   		COP(N746[TMP_dSourceOffset], N14[TMP_dDestOffset], TMP_dNumValues);
   	ELSIF (TMP_dSourceFile = 747) AND (TMP_dDestFile = 14) THEN
   		COP(N747[TMP_dSourceOffset], N14[TMP_dDestOffset], TMP_dNumValues);
   	ELSIF (TMP_dSourceFile = 748) AND (TMP_dDestFile = 14) THEN
   		COP(N748[TMP_dSourceOffset], N14[TMP_dDestOffset], TMP_dNumValues);
   	ELSIF (TMP_dSourceFile = 749) AND (TMP_dDestFile = 14) THEN
   		COP(N749[TMP_dSourceOffset], N14[TMP_dDestOffset], TMP_dNumValues);
   	ELSIF (TMP_dSourceFile = 750) AND (TMP_dDestFile = 14) THEN
   		COP(N750[TMP_dSourceOffset], N14[TMP_dDestOffset], TMP_dNumValues);
   	ELSIF (TMP_dSourceFile = 751) AND (TMP_dDestFile = 14) THEN
   		COP(N751[TMP_dSourceOffset], N14[TMP_dDestOffset], TMP_dNumValues);
   	ELSIF (TMP_dSourceFile = 752) AND (TMP_dDestFile = 14) THEN
   		COP(N752[TMP_dSourceOffset], N14[TMP_dDestOffset], TMP_dNumValues);
   	ELSIF (TMP_dSourceFile = 753) AND (TMP_dDestFile = 14) THEN
   		COP(N753[TMP_dSourceOffset], N14[TMP_dDestOffset], TMP_dNumValues);
   	ELSIF (TMP_dSourceFile = 754) AND (TMP_dDestFile = 14) THEN
   		COP(N754[TMP_dSourceOffset], N14[TMP_dDestOffset], TMP_dNumValues);
   	ELSIF (TMP_dSourceFile = 755) AND (TMP_dDestFile = 14) THEN
   		COP(N755[TMP_dSourceOffset], N14[TMP_dDestOffset], TMP_dNumValues);
   	ELSIF (TMP_dSourceFile = 756) AND (TMP_dDestFile = 14) THEN
   		COP(N756[TMP_dSourceOffset], N14[TMP_dDestOffset], TMP_dNumValues);
   	ELSIF (TMP_dSourceFile = 757) AND (TMP_dDestFile = 14) THEN
   		COP(N757[TMP_dSourceOffset], N14[TMP_dDestOffset], TMP_dNumValues);
   	ELSIF (TMP_dSourceFile = 758) AND (TMP_dDestFile = 14) THEN
   		COP(N758[TMP_dSourceOffset], N14[TMP_dDestOffset], TMP_dNumValues);
   	ELSIF (TMP_dSourceFile = 759) AND (TMP_dDestFile = 14) THEN
   		COP(N759[TMP_dSourceOffset], N14[TMP_dDestOffset], TMP_dNumValues);
   	ELSIF (TMP_dSourceFile = 760) AND (TMP_dDestFile = 14) THEN
   		COP(N760[TMP_dSourceOffset], N14[TMP_dDestOffset], TMP_dNumValues);
   	ELSIF (TMP_dSourceFile = 761) AND (TMP_dDestFile = 14) THEN
   		COP(N761[TMP_dSourceOffset], N14[TMP_dDestOffset], TMP_dNumValues);
   	ELSIF (TMP_dSourceFile = 762) AND (TMP_dDestFile = 14) THEN
   		COP(N762[TMP_dSourceOffset], N14[TMP_dDestOffset], TMP_dNumValues);
   	ELSIF (TMP_dSourceFile = 763) AND (TMP_dDestFile = 14) THEN
   		COP(N763[TMP_dSourceOffset], N14[TMP_dDestOffset], TMP_dNumValues);
   	ELSIF (TMP_dSourceFile = 764) AND (TMP_dDestFile = 14) THEN
   		COP(N764[TMP_dSourceOffset], N14[TMP_dDestOffset], TMP_dNumValues);
   	ELSIF (TMP_dSourceFile = 765) AND (TMP_dDestFile = 14) THEN
   		COP(N765[TMP_dSourceOffset], N14[TMP_dDestOffset], TMP_dNumValues);
   	ELSIF (TMP_dSourceFile = 766) AND (TMP_dDestFile = 14) THEN
   		COP(N766[TMP_dSourceOffset], N14[TMP_dDestOffset], TMP_dNumValues);
   	ELSIF (TMP_dSourceFile = 767) AND (TMP_dDestFile = 14) THEN
   		COP(N767[TMP_dSourceOffset], N14[TMP_dDestOffset], TMP_dNumValues);
   	ELSIF (TMP_dSourceFile = 768) AND (TMP_dDestFile = 14) THEN
   		COP(N768[TMP_dSourceOffset], N14[TMP_dDestOffset], TMP_dNumValues);
   	ELSIF (TMP_dSourceFile = 769) AND (TMP_dDestFile = 14) THEN
   		COP(N769[TMP_dSourceOffset], N14[TMP_dDestOffset], TMP_dNumValues);
   	ELSIF (TMP_dSourceFile = 770) AND (TMP_dDestFile = 14) THEN
   		COP(N770[TMP_dSourceOffset], N14[TMP_dDestOffset], TMP_dNumValues);
   	ELSIF (TMP_dSourceFile = 771) AND (TMP_dDestFile = 14) THEN
   		COP(N771[TMP_dSourceOffset], N14[TMP_dDestOffset], TMP_dNumValues);
   	ELSIF (TMP_dSourceFile = 772) AND (TMP_dDestFile = 14) THEN
   		COP(N772[TMP_dSourceOffset], N14[TMP_dDestOffset], TMP_dNumValues);
   	ELSIF (TMP_dSourceFile = 773) AND (TMP_dDestFile = 14) THEN
   		COP(N773[TMP_dSourceOffset], N14[TMP_dDestOffset], TMP_dNumValues);
   	ELSIF (TMP_dSourceFile = 774) AND (TMP_dDestFile = 14) THEN
   		COP(N774[TMP_dSourceOffset], N14[TMP_dDestOffset], TMP_dNumValues);
   	ELSIF (TMP_dSourceFile = 775) AND (TMP_dDestFile = 14) THEN
   		COP(N775[TMP_dSourceOffset], N14[TMP_dDestOffset], TMP_dNumValues);
   	ELSIF (TMP_dSourceFile = 776) AND (TMP_dDestFile = 14) THEN
   		COP(N776[TMP_dSourceOffset], N14[TMP_dDestOffset], TMP_dNumValues);
   	ELSIF (TMP_dSourceFile = 777) AND (TMP_dDestFile = 14) THEN
   		COP(N777[TMP_dSourceOffset], N14[TMP_dDestOffset], TMP_dNumValues);
   	ELSIF (TMP_dSourceFile = 778) AND (TMP_dDestFile = 14) THEN
   		COP(N778[TMP_dSourceOffset], N14[TMP_dDestOffset], TMP_dNumValues);
   	ELSIF (TMP_dSourceFile = 779) AND (TMP_dDestFile = 14) THEN
   		COP(N779[TMP_dSourceOffset], N14[TMP_dDestOffset], TMP_dNumValues);
   	ELSIF (TMP_dSourceFile = 780) AND (TMP_dDestFile = 14) THEN
   		COP(N780[TMP_dSourceOffset], N14[TMP_dDestOffset], TMP_dNumValues);
   	ELSIF (TMP_dSourceFile = 781) AND (TMP_dDestFile = 14) THEN
   		COP(N781[TMP_dSourceOffset], N14[TMP_dDestOffset], TMP_dNumValues);
   	ELSIF (TMP_dSourceFile = 782) AND (TMP_dDestFile = 14) THEN
   		COP(N782[TMP_dSourceOffset], N14[TMP_dDestOffset], TMP_dNumValues);
   	ELSIF (TMP_dSourceFile = 783) AND (TMP_dDestFile = 14) THEN
   		COP(N783[TMP_dSourceOffset], N14[TMP_dDestOffset], TMP_dNumValues);
   	ELSIF (TMP_dSourceFile = 784) AND (TMP_dDestFile = 14) THEN
   		COP(N784[TMP_dSourceOffset], N14[TMP_dDestOffset], TMP_dNumValues);
   	ELSIF (TMP_dSourceFile = 785) AND (TMP_dDestFile = 14) THEN
   		COP(N785[TMP_dSourceOffset], N14[TMP_dDestOffset], TMP_dNumValues);
   	ELSIF (TMP_dSourceFile = 786) AND (TMP_dDestFile = 14) THEN
   		COP(N786[TMP_dSourceOffset], N14[TMP_dDestOffset], TMP_dNumValues);
   	ELSIF (TMP_dSourceFile = 787) AND (TMP_dDestFile = 14) THEN
   		COP(N787[TMP_dSourceOffset], N14[TMP_dDestOffset], TMP_dNumValues);
   	ELSIF (TMP_dSourceFile = 788) AND (TMP_dDestFile = 14) THEN
   		COP(N788[TMP_dSourceOffset], N14[TMP_dDestOffset], TMP_dNumValues);
   	ELSIF (TMP_dSourceFile = 789) AND (TMP_dDestFile = 14) THEN
   		COP(N789[TMP_dSourceOffset], N14[TMP_dDestOffset], TMP_dNumValues);
   	ELSIF (TMP_dSourceFile = 790) AND (TMP_dDestFile = 14) THEN
   		COP(N790[TMP_dSourceOffset], N14[TMP_dDestOffset], TMP_dNumValues);
   	ELSIF (TMP_dSourceFile = 791) AND (TMP_dDestFile = 14) THEN
   		COP(N791[TMP_dSourceOffset], N14[TMP_dDestOffset], TMP_dNumValues);
   	ELSIF (TMP_dSourceFile = 792) AND (TMP_dDestFile = 14) THEN
   		COP(N792[TMP_dSourceOffset], N14[TMP_dDestOffset], TMP_dNumValues);
   	ELSIF (TMP_dSourceFile = 793) AND (TMP_dDestFile = 14) THEN
   		COP(N793[TMP_dSourceOffset], N14[TMP_dDestOffset], TMP_dNumValues);
   	ELSIF (TMP_dSourceFile = 794) AND (TMP_dDestFile = 14) THEN
   		COP(N794[TMP_dSourceOffset], N14[TMP_dDestOffset], TMP_dNumValues);
   	ELSIF (TMP_dSourceFile = 795) AND (TMP_dDestFile = 14) THEN
   		COP(N795[TMP_dSourceOffset], N14[TMP_dDestOffset], TMP_dNumValues);
   	ELSIF (TMP_dSourceFile = 796) AND (TMP_dDestFile = 14) THEN
   		COP(N796[TMP_dSourceOffset], N14[TMP_dDestOffset], TMP_dNumValues);
   	ELSIF (TMP_dSourceFile = 797) AND (TMP_dDestFile = 14) THEN
   		COP(N797[TMP_dSourceOffset], N14[TMP_dDestOffset], TMP_dNumValues);
   	ELSIF (TMP_dSourceFile = 798) AND (TMP_dDestFile = 14) THEN
   		COP(N798[TMP_dSourceOffset], N14[TMP_dDestOffset], TMP_dNumValues);
   	ELSIF (TMP_dSourceFile = 799) AND (TMP_dDestFile = 14) THEN
   		COP(N799[TMP_dSourceOffset], N14[TMP_dDestOffset], TMP_dNumValues);
   
   /*
   ////CAPIDINDEX N23
   	IF (TMP_dSourceFile = 23) AND (TMP_dDestFile = 601) THEN
   		COP(N23[TMP_dSourceOffset], N601[TMP_dDestOffset], TMP_dNumValues);
   	ELSIF (TMP_dSourceFile = 23) AND (TMP_dDestFile = 602) THEN
   		COP(N23[TMP_dSourceOffset], N602[TMP_dDestOffset], TMP_dNumValues);
   	ELSIF (TMP_dSourceFile = 23) AND (TMP_dDestFile = 603) THEN
   		COP(N23[TMP_dSourceOffset], N603[TMP_dDestOffset], TMP_dNumValues);
   	ELSIF (TMP_dSourceFile = 23) AND (TMP_dDestFile = 604) THEN
   		COP(N23[TMP_dSourceOffset], N604[TMP_dDestOffset], TMP_dNumValues);
   	ELSIF (TMP_dSourceFile = 23) AND (TMP_dDestFile = 605) THEN
   		COP(N23[TMP_dSourceOffset], N605[TMP_dDestOffset], TMP_dNumValues);
   	ELSIF (TMP_dSourceFile = 23) AND (TMP_dDestFile = 606) THEN
   		COP(N23[TMP_dSourceOffset], N606[TMP_dDestOffset], TMP_dNumValues);
   	ELSIF (TMP_dSourceFile = 23) AND (TMP_dDestFile = 607) THEN
   		COP(N23[TMP_dSourceOffset], N607[TMP_dDestOffset], TMP_dNumValues);
   	ELSIF (TMP_dSourceFile = 23) AND (TMP_dDestFile = 608) THEN
   		COP(N23[TMP_dSourceOffset], N608[TMP_dDestOffset], TMP_dNumValues);
   	ELSIF (TMP_dSourceFile = 23) AND (TMP_dDestFile = 609) THEN
   		COP(N23[TMP_dSourceOffset], N609[TMP_dDestOffset], TMP_dNumValues);
   	ELSIF (TMP_dSourceFile = 23) AND (TMP_dDestFile = 610) THEN
   		COP(N23[TMP_dSourceOffset], N610[TMP_dDestOffset], TMP_dNumValues);
   	ELSIF (TMP_dSourceFile = 23) AND (TMP_dDestFile = 611) THEN
   		COP(N23[TMP_dSourceOffset], N611[TMP_dDestOffset], TMP_dNumValues);
   	ELSIF (TMP_dSourceFile = 23) AND (TMP_dDestFile = 612) THEN
   		COP(N23[TMP_dSourceOffset], N612[TMP_dDestOffset], TMP_dNumValues);
   	ELSIF (TMP_dSourceFile = 23) AND (TMP_dDestFile = 613) THEN
   		COP(N23[TMP_dSourceOffset], N613[TMP_dDestOffset], TMP_dNumValues);
   	ELSIF (TMP_dSourceFile = 23) AND (TMP_dDestFile = 614) THEN
   		COP(N23[TMP_dSourceOffset], N614[TMP_dDestOffset], TMP_dNumValues);
   	ELSIF (TMP_dSourceFile = 23) AND (TMP_dDestFile = 615) THEN
   		COP(N23[TMP_dSourceOffset], N615[TMP_dDestOffset], TMP_dNumValues);
   	ELSIF (TMP_dSourceFile = 23) AND (TMP_dDestFile = 616) THEN
   		COP(N23[TMP_dSourceOffset], N616[TMP_dDestOffset], TMP_dNumValues);
   	ELSIF (TMP_dSourceFile = 23) AND (TMP_dDestFile = 617) THEN
   		COP(N23[TMP_dSourceOffset], N617[TMP_dDestOffset], TMP_dNumValues);
   	ELSIF (TMP_dSourceFile = 23) AND (TMP_dDestFile = 618) THEN
   		COP(N23[TMP_dSourceOffset], N618[TMP_dDestOffset], TMP_dNumValues);
   	ELSIF (TMP_dSourceFile = 23) AND (TMP_dDestFile = 619) THEN
   		COP(N23[TMP_dSourceOffset], N619[TMP_dDestOffset], TMP_dNumValues);
   	ELSIF (TMP_dSourceFile = 23) AND (TMP_dDestFile = 620) THEN
   		COP(N23[TMP_dSourceOffset], N620[TMP_dDestOffset], TMP_dNumValues);
   	ELSIF (TMP_dSourceFile = 23) AND (TMP_dDestFile = 621) THEN
   		COP(N23[TMP_dSourceOffset], N621[TMP_dDestOffset], TMP_dNumValues);
   	ELSIF (TMP_dSourceFile = 23) AND (TMP_dDestFile = 622) THEN
   		COP(N23[TMP_dSourceOffset], N622[TMP_dDestOffset], TMP_dNumValues);
   	ELSIF (TMP_dSourceFile = 23) AND (TMP_dDestFile = 623) THEN
   		COP(N23[TMP_dSourceOffset], N623[TMP_dDestOffset], TMP_dNumValues);
   	ELSIF (TMP_dSourceFile = 23) AND (TMP_dDestFile = 624) THEN
   		COP(N23[TMP_dSourceOffset], N624[TMP_dDestOffset], TMP_dNumValues);
   	ELSIF (TMP_dSourceFile = 23) AND (TMP_dDestFile = 625) THEN
   		COP(N23[TMP_dSourceOffset], N625[TMP_dDestOffset], TMP_dNumValues);
   	ELSIF (TMP_dSourceFile = 23) AND (TMP_dDestFile = 626) THEN
   		COP(N23[TMP_dSourceOffset], N626[TMP_dDestOffset], TMP_dNumValues);
   	ELSIF (TMP_dSourceFile = 23) AND (TMP_dDestFile = 627) THEN
   		COP(N23[TMP_dSourceOffset], N627[TMP_dDestOffset], TMP_dNumValues);
   	ELSIF (TMP_dSourceFile = 23) AND (TMP_dDestFile = 628) THEN
   		COP(N23[TMP_dSourceOffset], N628[TMP_dDestOffset], TMP_dNumValues);
   	ELSIF (TMP_dSourceFile = 23) AND (TMP_dDestFile = 629) THEN
   		COP(N23[TMP_dSourceOffset], N629[TMP_dDestOffset], TMP_dNumValues);
   	ELSIF (TMP_dSourceFile = 23) AND (TMP_dDestFile = 630) THEN
   		COP(N23[TMP_dSourceOffset], N630[TMP_dDestOffset], TMP_dNumValues);
   	ELSIF (TMP_dSourceFile = 23) AND (TMP_dDestFile = 631) THEN
   		COP(N23[TMP_dSourceOffset], N631[TMP_dDestOffset], TMP_dNumValues);
   	ELSIF (TMP_dSourceFile = 23) AND (TMP_dDestFile = 632) THEN
   		COP(N23[TMP_dSourceOffset], N632[TMP_dDestOffset], TMP_dNumValues);
   	ELSIF (TMP_dSourceFile = 23) AND (TMP_dDestFile = 633) THEN
   		COP(N23[TMP_dSourceOffset], N633[TMP_dDestOffset], TMP_dNumValues);
   	ELSIF (TMP_dSourceFile = 23) AND (TMP_dDestFile = 634) THEN
   		COP(N23[TMP_dSourceOffset], N634[TMP_dDestOffset], TMP_dNumValues);
   	ELSIF (TMP_dSourceFile = 23) AND (TMP_dDestFile = 635) THEN
   		COP(N23[TMP_dSourceOffset], N635[TMP_dDestOffset], TMP_dNumValues);
   	ELSIF (TMP_dSourceFile = 23) AND (TMP_dDestFile = 636) THEN
   		COP(N23[TMP_dSourceOffset], N636[TMP_dDestOffset], TMP_dNumValues);
   	ELSIF (TMP_dSourceFile = 23) AND (TMP_dDestFile = 637) THEN
   		COP(N23[TMP_dSourceOffset], N637[TMP_dDestOffset], TMP_dNumValues);
   	ELSIF (TMP_dSourceFile = 23) AND (TMP_dDestFile = 638) THEN
   		COP(N23[TMP_dSourceOffset], N638[TMP_dDestOffset], TMP_dNumValues);
   	ELSIF (TMP_dSourceFile = 23) AND (TMP_dDestFile = 639) THEN
   		COP(N23[TMP_dSourceOffset], N639[TMP_dDestOffset], TMP_dNumValues);
   	ELSIF (TMP_dSourceFile = 23) AND (TMP_dDestFile = 640) THEN
   		COP(N23[TMP_dSourceOffset], N640[TMP_dDestOffset], TMP_dNumValues);
   	ELSIF (TMP_dSourceFile = 23) AND (TMP_dDestFile = 641) THEN
   		COP(N23[TMP_dSourceOffset], N641[TMP_dDestOffset], TMP_dNumValues);
   	ELSIF (TMP_dSourceFile = 23) AND (TMP_dDestFile = 642) THEN
   		COP(N23[TMP_dSourceOffset], N642[TMP_dDestOffset], TMP_dNumValues);
   	ELSIF (TMP_dSourceFile = 23) AND (TMP_dDestFile = 643) THEN
   		COP(N23[TMP_dSourceOffset], N643[TMP_dDestOffset], TMP_dNumValues);
   	ELSIF (TMP_dSourceFile = 23) AND (TMP_dDestFile = 644) THEN
   		COP(N23[TMP_dSourceOffset], N644[TMP_dDestOffset], TMP_dNumValues);
   	ELSIF (TMP_dSourceFile = 23) AND (TMP_dDestFile = 645) THEN
   		COP(N23[TMP_dSourceOffset], N645[TMP_dDestOffset], TMP_dNumValues);
   	ELSIF (TMP_dSourceFile = 23) AND (TMP_dDestFile = 646) THEN
   		COP(N23[TMP_dSourceOffset], N646[TMP_dDestOffset], TMP_dNumValues);
   	ELSIF (TMP_dSourceFile = 23) AND (TMP_dDestFile = 647) THEN
   		COP(N23[TMP_dSourceOffset], N647[TMP_dDestOffset], TMP_dNumValues);
   	ELSIF (TMP_dSourceFile = 23) AND (TMP_dDestFile = 648) THEN
   		COP(N23[TMP_dSourceOffset], N648[TMP_dDestOffset], TMP_dNumValues);
   	ELSIF (TMP_dSourceFile = 23) AND (TMP_dDestFile = 649) THEN
   		COP(N23[TMP_dSourceOffset], N649[TMP_dDestOffset], TMP_dNumValues);
   	ELSIF (TMP_dSourceFile = 23) AND (TMP_dDestFile = 650) THEN
   		COP(N23[TMP_dSourceOffset], N650[TMP_dDestOffset], TMP_dNumValues);
   	ELSIF (TMP_dSourceFile = 23) AND (TMP_dDestFile = 651) THEN
   		COP(N23[TMP_dSourceOffset], N651[TMP_dDestOffset], TMP_dNumValues);
   	ELSIF (TMP_dSourceFile = 23) AND (TMP_dDestFile = 652) THEN
   		COP(N23[TMP_dSourceOffset], N652[TMP_dDestOffset], TMP_dNumValues);
   	ELSIF (TMP_dSourceFile = 23) AND (TMP_dDestFile = 653) THEN
   		COP(N23[TMP_dSourceOffset], N653[TMP_dDestOffset], TMP_dNumValues);
   	ELSIF (TMP_dSourceFile = 23) AND (TMP_dDestFile = 654) THEN
   		COP(N23[TMP_dSourceOffset], N654[TMP_dDestOffset], TMP_dNumValues);
   	ELSIF (TMP_dSourceFile = 23) AND (TMP_dDestFile = 655) THEN
   		COP(N23[TMP_dSourceOffset], N655[TMP_dDestOffset], TMP_dNumValues);
   	ELSIF (TMP_dSourceFile = 23) AND (TMP_dDestFile = 656) THEN
   		COP(N23[TMP_dSourceOffset], N656[TMP_dDestOffset], TMP_dNumValues);
   	ELSIF (TMP_dSourceFile = 23) AND (TMP_dDestFile = 657) THEN
   		COP(N23[TMP_dSourceOffset], N657[TMP_dDestOffset], TMP_dNumValues);
   	ELSIF (TMP_dSourceFile = 23) AND (TMP_dDestFile = 658) THEN
   		COP(N23[TMP_dSourceOffset], N658[TMP_dDestOffset], TMP_dNumValues);
   	ELSIF (TMP_dSourceFile = 23) AND (TMP_dDestFile = 659) THEN
   		COP(N23[TMP_dSourceOffset], N659[TMP_dDestOffset], TMP_dNumValues);
   	ELSIF (TMP_dSourceFile = 23) AND (TMP_dDestFile = 660) THEN
   		COP(N23[TMP_dSourceOffset], N660[TMP_dDestOffset], TMP_dNumValues);
   	ELSIF (TMP_dSourceFile = 23) AND (TMP_dDestFile = 661) THEN
   		COP(N23[TMP_dSourceOffset], N661[TMP_dDestOffset], TMP_dNumValues);
   	ELSIF (TMP_dSourceFile = 23) AND (TMP_dDestFile = 662) THEN
   		COP(N23[TMP_dSourceOffset], N662[TMP_dDestOffset], TMP_dNumValues);
   	ELSIF (TMP_dSourceFile = 23) AND (TMP_dDestFile = 663) THEN
   		COP(N23[TMP_dSourceOffset], N663[TMP_dDestOffset], TMP_dNumValues);
   	ELSIF (TMP_dSourceFile = 23) AND (TMP_dDestFile = 664) THEN
   		COP(N23[TMP_dSourceOffset], N664[TMP_dDestOffset], TMP_dNumValues);
   	ELSIF (TMP_dSourceFile = 23) AND (TMP_dDestFile = 665) THEN
   		COP(N23[TMP_dSourceOffset], N665[TMP_dDestOffset], TMP_dNumValues);
   	ELSIF (TMP_dSourceFile = 23) AND (TMP_dDestFile = 666) THEN
   		COP(N23[TMP_dSourceOffset], N666[TMP_dDestOffset], TMP_dNumValues);
   	ELSIF (TMP_dSourceFile = 23) AND (TMP_dDestFile = 667) THEN
   		COP(N23[TMP_dSourceOffset], N667[TMP_dDestOffset], TMP_dNumValues);
   	ELSIF (TMP_dSourceFile = 23) AND (TMP_dDestFile = 668) THEN
   		COP(N23[TMP_dSourceOffset], N668[TMP_dDestOffset], TMP_dNumValues);
   	ELSIF (TMP_dSourceFile = 23) AND (TMP_dDestFile = 669) THEN
   		COP(N23[TMP_dSourceOffset], N669[TMP_dDestOffset], TMP_dNumValues);
   	ELSIF (TMP_dSourceFile = 23) AND (TMP_dDestFile = 670) THEN
   		COP(N23[TMP_dSourceOffset], N670[TMP_dDestOffset], TMP_dNumValues);
   	ELSIF (TMP_dSourceFile = 23) AND (TMP_dDestFile = 671) THEN
   		COP(N23[TMP_dSourceOffset], N671[TMP_dDestOffset], TMP_dNumValues);
   	ELSIF (TMP_dSourceFile = 23) AND (TMP_dDestFile = 672) THEN
   		COP(N23[TMP_dSourceOffset], N672[TMP_dDestOffset], TMP_dNumValues);
   	ELSIF (TMP_dSourceFile = 23) AND (TMP_dDestFile = 673) THEN
   		COP(N23[TMP_dSourceOffset], N673[TMP_dDestOffset], TMP_dNumValues);
   	ELSIF (TMP_dSourceFile = 23) AND (TMP_dDestFile = 674) THEN
   		COP(N23[TMP_dSourceOffset], N674[TMP_dDestOffset], TMP_dNumValues);
   	ELSIF (TMP_dSourceFile = 23) AND (TMP_dDestFile = 675) THEN
   		COP(N23[TMP_dSourceOffset], N675[TMP_dDestOffset], TMP_dNumValues);
   	ELSIF (TMP_dSourceFile = 23) AND (TMP_dDestFile = 676) THEN
   		COP(N23[TMP_dSourceOffset], N676[TMP_dDestOffset], TMP_dNumValues);
   	ELSIF (TMP_dSourceFile = 23) AND (TMP_dDestFile = 677) THEN
   		COP(N23[TMP_dSourceOffset], N677[TMP_dDestOffset], TMP_dNumValues);
   	ELSIF (TMP_dSourceFile = 23) AND (TMP_dDestFile = 678) THEN
   		COP(N23[TMP_dSourceOffset], N678[TMP_dDestOffset], TMP_dNumValues);
   	ELSIF (TMP_dSourceFile = 23) AND (TMP_dDestFile = 679) THEN
   		COP(N23[TMP_dSourceOffset], N679[TMP_dDestOffset], TMP_dNumValues);
   	ELSIF (TMP_dSourceFile = 23) AND (TMP_dDestFile = 680) THEN
   		COP(N23[TMP_dSourceOffset], N680[TMP_dDestOffset], TMP_dNumValues);
   	ELSIF (TMP_dSourceFile = 23) AND (TMP_dDestFile = 681) THEN
   		COP(N23[TMP_dSourceOffset], N681[TMP_dDestOffset], TMP_dNumValues);
   	ELSIF (TMP_dSourceFile = 23) AND (TMP_dDestFile = 682) THEN
   		COP(N23[TMP_dSourceOffset], N682[TMP_dDestOffset], TMP_dNumValues);
   	ELSIF (TMP_dSourceFile = 23) AND (TMP_dDestFile = 683) THEN
   		COP(N23[TMP_dSourceOffset], N683[TMP_dDestOffset], TMP_dNumValues);
   	ELSIF (TMP_dSourceFile = 23) AND (TMP_dDestFile = 684) THEN
   		COP(N23[TMP_dSourceOffset], N684[TMP_dDestOffset], TMP_dNumValues);
   	ELSIF (TMP_dSourceFile = 23) AND (TMP_dDestFile = 685) THEN
   		COP(N23[TMP_dSourceOffset], N685[TMP_dDestOffset], TMP_dNumValues);
   	ELSIF (TMP_dSourceFile = 23) AND (TMP_dDestFile = 686) THEN
   		COP(N23[TMP_dSourceOffset], N686[TMP_dDestOffset], TMP_dNumValues);
   	ELSIF (TMP_dSourceFile = 23) AND (TMP_dDestFile = 687) THEN
   		COP(N23[TMP_dSourceOffset], N687[TMP_dDestOffset], TMP_dNumValues);
   	ELSIF (TMP_dSourceFile = 23) AND (TMP_dDestFile = 688) THEN
   		COP(N23[TMP_dSourceOffset], N688[TMP_dDestOffset], TMP_dNumValues);
   	ELSIF (TMP_dSourceFile = 23) AND (TMP_dDestFile = 689) THEN
   		COP(N23[TMP_dSourceOffset], N689[TMP_dDestOffset], TMP_dNumValues);
   	ELSIF (TMP_dSourceFile = 23) AND (TMP_dDestFile = 690) THEN
   		COP(N23[TMP_dSourceOffset], N690[TMP_dDestOffset], TMP_dNumValues);
   	ELSIF (TMP_dSourceFile = 23) AND (TMP_dDestFile = 691) THEN
   		COP(N23[TMP_dSourceOffset], N691[TMP_dDestOffset], TMP_dNumValues);
   	ELSIF (TMP_dSourceFile = 23) AND (TMP_dDestFile = 692) THEN
   		COP(N23[TMP_dSourceOffset], N692[TMP_dDestOffset], TMP_dNumValues);
   	ELSIF (TMP_dSourceFile = 23) AND (TMP_dDestFile = 693) THEN
   		COP(N23[TMP_dSourceOffset], N693[TMP_dDestOffset], TMP_dNumValues);
   	ELSIF (TMP_dSourceFile = 23) AND (TMP_dDestFile = 694) THEN
   		COP(N23[TMP_dSourceOffset], N694[TMP_dDestOffset], TMP_dNumValues);
   	ELSIF (TMP_dSourceFile = 23) AND (TMP_dDestFile = 695) THEN
   		COP(N23[TMP_dSourceOffset], N695[TMP_dDestOffset], TMP_dNumValues);
   	ELSIF (TMP_dSourceFile = 23) AND (TMP_dDestFile = 696) THEN
   		COP(N23[TMP_dSourceOffset], N696[TMP_dDestOffset], TMP_dNumValues);
   	ELSIF (TMP_dSourceFile = 23) AND (TMP_dDestFile = 697) THEN
   		COP(N23[TMP_dSourceOffset], N697[TMP_dDestOffset], TMP_dNumValues);
   	ELSIF (TMP_dSourceFile = 23) AND (TMP_dDestFile = 698) THEN
   		COP(N23[TMP_dSourceOffset], N698[TMP_dDestOffset], TMP_dNumValues);
   	ELSIF (TMP_dSourceFile = 23) AND (TMP_dDestFile = 699) THEN
   		COP(N23[TMP_dSourceOffset], N699[TMP_dDestOffset], TMP_dNumValues);
   	ELSIF (TMP_dSourceFile = 23) AND (TMP_dDestFile = 700) THEN
   		COP(N23[TMP_dSourceOffset], N700[TMP_dDestOffset], TMP_dNumValues);
   	ELSIF (TMP_dSourceFile = 23) AND (TMP_dDestFile = 701) THEN
   		COP(N23[TMP_dSourceOffset], N701[TMP_dDestOffset], TMP_dNumValues);
   	ELSIF (TMP_dSourceFile = 23) AND (TMP_dDestFile = 702) THEN
   		COP(N23[TMP_dSourceOffset], N702[TMP_dDestOffset], TMP_dNumValues);
   	ELSIF (TMP_dSourceFile = 23) AND (TMP_dDestFile = 703) THEN
   		COP(N23[TMP_dSourceOffset], N703[TMP_dDestOffset], TMP_dNumValues);
   	ELSIF (TMP_dSourceFile = 23) AND (TMP_dDestFile = 704) THEN
   		COP(N23[TMP_dSourceOffset], N704[TMP_dDestOffset], TMP_dNumValues);
   	ELSIF (TMP_dSourceFile = 23) AND (TMP_dDestFile = 705) THEN
   		COP(N23[TMP_dSourceOffset], N705[TMP_dDestOffset], TMP_dNumValues);
   	ELSIF (TMP_dSourceFile = 23) AND (TMP_dDestFile = 706) THEN
   		COP(N23[TMP_dSourceOffset], N706[TMP_dDestOffset], TMP_dNumValues);
   	ELSIF (TMP_dSourceFile = 23) AND (TMP_dDestFile = 707) THEN
   		COP(N23[TMP_dSourceOffset], N707[TMP_dDestOffset], TMP_dNumValues);
   	ELSIF (TMP_dSourceFile = 23) AND (TMP_dDestFile = 708) THEN
   		COP(N23[TMP_dSourceOffset], N708[TMP_dDestOffset], TMP_dNumValues);
   	ELSIF (TMP_dSourceFile = 23) AND (TMP_dDestFile = 709) THEN
   		COP(N23[TMP_dSourceOffset], N709[TMP_dDestOffset], TMP_dNumValues);
   	ELSIF (TMP_dSourceFile = 23) AND (TMP_dDestFile = 710) THEN
   		COP(N23[TMP_dSourceOffset], N710[TMP_dDestOffset], TMP_dNumValues);
   	ELSIF (TMP_dSourceFile = 23) AND (TMP_dDestFile = 711) THEN
   		COP(N23[TMP_dSourceOffset], N711[TMP_dDestOffset], TMP_dNumValues);
   	ELSIF (TMP_dSourceFile = 23) AND (TMP_dDestFile = 712) THEN
   		COP(N23[TMP_dSourceOffset], N712[TMP_dDestOffset], TMP_dNumValues);
   	ELSIF (TMP_dSourceFile = 23) AND (TMP_dDestFile = 713) THEN
   		COP(N23[TMP_dSourceOffset], N713[TMP_dDestOffset], TMP_dNumValues);
   	ELSIF (TMP_dSourceFile = 23) AND (TMP_dDestFile = 714) THEN
   		COP(N23[TMP_dSourceOffset], N714[TMP_dDestOffset], TMP_dNumValues);
   	ELSIF (TMP_dSourceFile = 23) AND (TMP_dDestFile = 715) THEN
   		COP(N23[TMP_dSourceOffset], N715[TMP_dDestOffset], TMP_dNumValues);
   	ELSIF (TMP_dSourceFile = 23) AND (TMP_dDestFile = 716) THEN
   		COP(N23[TMP_dSourceOffset], N716[TMP_dDestOffset], TMP_dNumValues);
   	ELSIF (TMP_dSourceFile = 23) AND (TMP_dDestFile = 717) THEN
   		COP(N23[TMP_dSourceOffset], N717[TMP_dDestOffset], TMP_dNumValues);
   	ELSIF (TMP_dSourceFile = 23) AND (TMP_dDestFile = 718) THEN
   		COP(N23[TMP_dSourceOffset], N718[TMP_dDestOffset], TMP_dNumValues);
   	ELSIF (TMP_dSourceFile = 23) AND (TMP_dDestFile = 719) THEN
   		COP(N23[TMP_dSourceOffset], N719[TMP_dDestOffset], TMP_dNumValues);
   	ELSIF (TMP_dSourceFile = 23) AND (TMP_dDestFile = 720) THEN
   		COP(N23[TMP_dSourceOffset], N720[TMP_dDestOffset], TMP_dNumValues);
   	ELSIF (TMP_dSourceFile = 23) AND (TMP_dDestFile = 721) THEN
   		COP(N23[TMP_dSourceOffset], N721[TMP_dDestOffset], TMP_dNumValues);
   	ELSIF (TMP_dSourceFile = 23) AND (TMP_dDestFile = 722) THEN
   		COP(N23[TMP_dSourceOffset], N722[TMP_dDestOffset], TMP_dNumValues);
   	ELSIF (TMP_dSourceFile = 23) AND (TMP_dDestFile = 723) THEN
   		COP(N23[TMP_dSourceOffset], N723[TMP_dDestOffset], TMP_dNumValues);
   	ELSIF (TMP_dSourceFile = 23) AND (TMP_dDestFile = 724) THEN
   		COP(N23[TMP_dSourceOffset], N724[TMP_dDestOffset], TMP_dNumValues);
   	ELSIF (TMP_dSourceFile = 23) AND (TMP_dDestFile = 725) THEN
   		COP(N23[TMP_dSourceOffset], N725[TMP_dDestOffset], TMP_dNumValues);
   	ELSIF (TMP_dSourceFile = 23) AND (TMP_dDestFile = 726) THEN
   		COP(N23[TMP_dSourceOffset], N726[TMP_dDestOffset], TMP_dNumValues);
   	ELSIF (TMP_dSourceFile = 23) AND (TMP_dDestFile = 727) THEN
   		COP(N23[TMP_dSourceOffset], N727[TMP_dDestOffset], TMP_dNumValues);
   	ELSIF (TMP_dSourceFile = 23) AND (TMP_dDestFile = 728) THEN
   		COP(N23[TMP_dSourceOffset], N728[TMP_dDestOffset], TMP_dNumValues);
   	ELSIF (TMP_dSourceFile = 23) AND (TMP_dDestFile = 729) THEN
   		COP(N23[TMP_dSourceOffset], N729[TMP_dDestOffset], TMP_dNumValues);
   	ELSIF (TMP_dSourceFile = 23) AND (TMP_dDestFile = 730) THEN
   		COP(N23[TMP_dSourceOffset], N730[TMP_dDestOffset], TMP_dNumValues);
   	ELSIF (TMP_dSourceFile = 23) AND (TMP_dDestFile = 731) THEN
   		COP(N23[TMP_dSourceOffset], N731[TMP_dDestOffset], TMP_dNumValues);
   	ELSIF (TMP_dSourceFile = 23) AND (TMP_dDestFile = 732) THEN
   		COP(N23[TMP_dSourceOffset], N732[TMP_dDestOffset], TMP_dNumValues);
   	ELSIF (TMP_dSourceFile = 23) AND (TMP_dDestFile = 733) THEN
   		COP(N23[TMP_dSourceOffset], N733[TMP_dDestOffset], TMP_dNumValues);
   	ELSIF (TMP_dSourceFile = 23) AND (TMP_dDestFile = 734) THEN
   		COP(N23[TMP_dSourceOffset], N734[TMP_dDestOffset], TMP_dNumValues);
   	ELSIF (TMP_dSourceFile = 23) AND (TMP_dDestFile = 735) THEN
   		COP(N23[TMP_dSourceOffset], N735[TMP_dDestOffset], TMP_dNumValues);
   	ELSIF (TMP_dSourceFile = 23) AND (TMP_dDestFile = 736) THEN
   		COP(N23[TMP_dSourceOffset], N736[TMP_dDestOffset], TMP_dNumValues);
   	ELSIF (TMP_dSourceFile = 23) AND (TMP_dDestFile = 737) THEN
   		COP(N23[TMP_dSourceOffset], N737[TMP_dDestOffset], TMP_dNumValues);
   	ELSIF (TMP_dSourceFile = 23) AND (TMP_dDestFile = 738) THEN
   		COP(N23[TMP_dSourceOffset], N738[TMP_dDestOffset], TMP_dNumValues);
   	ELSIF (TMP_dSourceFile = 23) AND (TMP_dDestFile = 739) THEN
   		COP(N23[TMP_dSourceOffset], N739[TMP_dDestOffset], TMP_dNumValues);
   	ELSIF (TMP_dSourceFile = 23) AND (TMP_dDestFile = 740) THEN
   		COP(N23[TMP_dSourceOffset], N740[TMP_dDestOffset], TMP_dNumValues);
   	ELSIF (TMP_dSourceFile = 23) AND (TMP_dDestFile = 741) THEN
   		COP(N23[TMP_dSourceOffset], N741[TMP_dDestOffset], TMP_dNumValues);
   	ELSIF (TMP_dSourceFile = 23) AND (TMP_dDestFile = 742) THEN
   		COP(N23[TMP_dSourceOffset], N742[TMP_dDestOffset], TMP_dNumValues);
   	ELSIF (TMP_dSourceFile = 23) AND (TMP_dDestFile = 743) THEN
   		COP(N23[TMP_dSourceOffset], N743[TMP_dDestOffset], TMP_dNumValues);
   	ELSIF (TMP_dSourceFile = 23) AND (TMP_dDestFile = 744) THEN
   		COP(N23[TMP_dSourceOffset], N744[TMP_dDestOffset], TMP_dNumValues);
   	ELSIF (TMP_dSourceFile = 23) AND (TMP_dDestFile = 745) THEN
   		COP(N23[TMP_dSourceOffset], N745[TMP_dDestOffset], TMP_dNumValues);
   	ELSIF (TMP_dSourceFile = 23) AND (TMP_dDestFile = 746) THEN
   		COP(N23[TMP_dSourceOffset], N746[TMP_dDestOffset], TMP_dNumValues);
   	ELSIF (TMP_dSourceFile = 23) AND (TMP_dDestFile = 747) THEN
   		COP(N23[TMP_dSourceOffset], N747[TMP_dDestOffset], TMP_dNumValues);
   	ELSIF (TMP_dSourceFile = 23) AND (TMP_dDestFile = 748) THEN
   		COP(N23[TMP_dSourceOffset], N748[TMP_dDestOffset], TMP_dNumValues);
   	ELSIF (TMP_dSourceFile = 23) AND (TMP_dDestFile = 749) THEN
   		COP(N23[TMP_dSourceOffset], N749[TMP_dDestOffset], TMP_dNumValues);
   	ELSIF (TMP_dSourceFile = 23) AND (TMP_dDestFile = 750) THEN
   		COP(N23[TMP_dSourceOffset], N750[TMP_dDestOffset], TMP_dNumValues);
   	ELSIF (TMP_dSourceFile = 23) AND (TMP_dDestFile = 751) THEN
   		COP(N23[TMP_dSourceOffset], N751[TMP_dDestOffset], TMP_dNumValues);
   	ELSIF (TMP_dSourceFile = 23) AND (TMP_dDestFile = 752) THEN
   		COP(N23[TMP_dSourceOffset], N752[TMP_dDestOffset], TMP_dNumValues);
   	ELSIF (TMP_dSourceFile = 23) AND (TMP_dDestFile = 753) THEN
   		COP(N23[TMP_dSourceOffset], N753[TMP_dDestOffset], TMP_dNumValues);
   	ELSIF (TMP_dSourceFile = 23) AND (TMP_dDestFile = 754) THEN
   		COP(N23[TMP_dSourceOffset], N754[TMP_dDestOffset], TMP_dNumValues);
   	ELSIF (TMP_dSourceFile = 23) AND (TMP_dDestFile = 755) THEN
   		COP(N23[TMP_dSourceOffset], N755[TMP_dDestOffset], TMP_dNumValues);
   	ELSIF (TMP_dSourceFile = 23) AND (TMP_dDestFile = 756) THEN
   		COP(N23[TMP_dSourceOffset], N756[TMP_dDestOffset], TMP_dNumValues);
   	ELSIF (TMP_dSourceFile = 23) AND (TMP_dDestFile = 757) THEN
   		COP(N23[TMP_dSourceOffset], N757[TMP_dDestOffset], TMP_dNumValues);
   	ELSIF (TMP_dSourceFile = 23) AND (TMP_dDestFile = 758) THEN
   		COP(N23[TMP_dSourceOffset], N758[TMP_dDestOffset], TMP_dNumValues);
   	ELSIF (TMP_dSourceFile = 23) AND (TMP_dDestFile = 759) THEN
   		COP(N23[TMP_dSourceOffset], N759[TMP_dDestOffset], TMP_dNumValues);
   	ELSIF (TMP_dSourceFile = 23) AND (TMP_dDestFile = 760) THEN
   		COP(N23[TMP_dSourceOffset], N760[TMP_dDestOffset], TMP_dNumValues);
   	ELSIF (TMP_dSourceFile = 23) AND (TMP_dDestFile = 761) THEN
   		COP(N23[TMP_dSourceOffset], N761[TMP_dDestOffset], TMP_dNumValues);
   	ELSIF (TMP_dSourceFile = 23) AND (TMP_dDestFile = 762) THEN
   		COP(N23[TMP_dSourceOffset], N762[TMP_dDestOffset], TMP_dNumValues);
   	ELSIF (TMP_dSourceFile = 23) AND (TMP_dDestFile = 763) THEN
   		COP(N23[TMP_dSourceOffset], N763[TMP_dDestOffset], TMP_dNumValues);
   	ELSIF (TMP_dSourceFile = 23) AND (TMP_dDestFile = 764) THEN
   		COP(N23[TMP_dSourceOffset], N764[TMP_dDestOffset], TMP_dNumValues);
   	ELSIF (TMP_dSourceFile = 23) AND (TMP_dDestFile = 765) THEN
   		COP(N23[TMP_dSourceOffset], N765[TMP_dDestOffset], TMP_dNumValues);
   	ELSIF (TMP_dSourceFile = 23) AND (TMP_dDestFile = 766) THEN
   		COP(N23[TMP_dSourceOffset], N766[TMP_dDestOffset], TMP_dNumValues);
   	ELSIF (TMP_dSourceFile = 23) AND (TMP_dDestFile = 767) THEN
   		COP(N23[TMP_dSourceOffset], N767[TMP_dDestOffset], TMP_dNumValues);
   	ELSIF (TMP_dSourceFile = 23) AND (TMP_dDestFile = 768) THEN
   		COP(N23[TMP_dSourceOffset], N768[TMP_dDestOffset], TMP_dNumValues);
   	ELSIF (TMP_dSourceFile = 23) AND (TMP_dDestFile = 769) THEN
   		COP(N23[TMP_dSourceOffset], N769[TMP_dDestOffset], TMP_dNumValues);
   	ELSIF (TMP_dSourceFile = 23) AND (TMP_dDestFile = 770) THEN
   		COP(N23[TMP_dSourceOffset], N770[TMP_dDestOffset], TMP_dNumValues);
   	ELSIF (TMP_dSourceFile = 23) AND (TMP_dDestFile = 771) THEN
   		COP(N23[TMP_dSourceOffset], N771[TMP_dDestOffset], TMP_dNumValues);
   	ELSIF (TMP_dSourceFile = 23) AND (TMP_dDestFile = 772) THEN
   		COP(N23[TMP_dSourceOffset], N772[TMP_dDestOffset], TMP_dNumValues);
   	ELSIF (TMP_dSourceFile = 23) AND (TMP_dDestFile = 773) THEN
   		COP(N23[TMP_dSourceOffset], N773[TMP_dDestOffset], TMP_dNumValues);
   	ELSIF (TMP_dSourceFile = 23) AND (TMP_dDestFile = 774) THEN
   		COP(N23[TMP_dSourceOffset], N774[TMP_dDestOffset], TMP_dNumValues);
   	ELSIF (TMP_dSourceFile = 23) AND (TMP_dDestFile = 775) THEN
   		COP(N23[TMP_dSourceOffset], N775[TMP_dDestOffset], TMP_dNumValues);
   	ELSIF (TMP_dSourceFile = 23) AND (TMP_dDestFile = 776) THEN
   		COP(N23[TMP_dSourceOffset], N776[TMP_dDestOffset], TMP_dNumValues);
   	ELSIF (TMP_dSourceFile = 23) AND (TMP_dDestFile = 777) THEN
   		COP(N23[TMP_dSourceOffset], N777[TMP_dDestOffset], TMP_dNumValues);
   	ELSIF (TMP_dSourceFile = 23) AND (TMP_dDestFile = 778) THEN
   		COP(N23[TMP_dSourceOffset], N778[TMP_dDestOffset], TMP_dNumValues);
   	ELSIF (TMP_dSourceFile = 23) AND (TMP_dDestFile = 779) THEN
   		COP(N23[TMP_dSourceOffset], N779[TMP_dDestOffset], TMP_dNumValues);
   	ELSIF (TMP_dSourceFile = 23) AND (TMP_dDestFile = 780) THEN
   		COP(N23[TMP_dSourceOffset], N780[TMP_dDestOffset], TMP_dNumValues);
   	ELSIF (TMP_dSourceFile = 23) AND (TMP_dDestFile = 781) THEN
   		COP(N23[TMP_dSourceOffset], N781[TMP_dDestOffset], TMP_dNumValues);
   	ELSIF (TMP_dSourceFile = 23) AND (TMP_dDestFile = 782) THEN
   		COP(N23[TMP_dSourceOffset], N782[TMP_dDestOffset], TMP_dNumValues);
   	ELSIF (TMP_dSourceFile = 23) AND (TMP_dDestFile = 783) THEN
   		COP(N23[TMP_dSourceOffset], N783[TMP_dDestOffset], TMP_dNumValues);
   	ELSIF (TMP_dSourceFile = 23) AND (TMP_dDestFile = 784) THEN
   		COP(N23[TMP_dSourceOffset], N784[TMP_dDestOffset], TMP_dNumValues);
   	ELSIF (TMP_dSourceFile = 23) AND (TMP_dDestFile = 785) THEN
   		COP(N23[TMP_dSourceOffset], N785[TMP_dDestOffset], TMP_dNumValues);
   	ELSIF (TMP_dSourceFile = 23) AND (TMP_dDestFile = 786) THEN
   		COP(N23[TMP_dSourceOffset], N786[TMP_dDestOffset], TMP_dNumValues);
   	ELSIF (TMP_dSourceFile = 23) AND (TMP_dDestFile = 787) THEN
   		COP(N23[TMP_dSourceOffset], N787[TMP_dDestOffset], TMP_dNumValues);
   	ELSIF (TMP_dSourceFile = 23) AND (TMP_dDestFile = 788) THEN
   		COP(N23[TMP_dSourceOffset], N788[TMP_dDestOffset], TMP_dNumValues);
   	ELSIF (TMP_dSourceFile = 23) AND (TMP_dDestFile = 789) THEN
   		COP(N23[TMP_dSourceOffset], N789[TMP_dDestOffset], TMP_dNumValues);
   	ELSIF (TMP_dSourceFile = 23) AND (TMP_dDestFile = 790) THEN
   		COP(N23[TMP_dSourceOffset], N790[TMP_dDestOffset], TMP_dNumValues);
   	ELSIF (TMP_dSourceFile = 23) AND (TMP_dDestFile = 791) THEN
   		COP(N23[TMP_dSourceOffset], N791[TMP_dDestOffset], TMP_dNumValues);
   	ELSIF (TMP_dSourceFile = 23) AND (TMP_dDestFile = 792) THEN
   		COP(N23[TMP_dSourceOffset], N792[TMP_dDestOffset], TMP_dNumValues);
   	ELSIF (TMP_dSourceFile = 23) AND (TMP_dDestFile = 793) THEN
   		COP(N23[TMP_dSourceOffset], N793[TMP_dDestOffset], TMP_dNumValues);
   	ELSIF (TMP_dSourceFile = 23) AND (TMP_dDestFile = 794) THEN
   		COP(N23[TMP_dSourceOffset], N794[TMP_dDestOffset], TMP_dNumValues);
   	ELSIF (TMP_dSourceFile = 23) AND (TMP_dDestFile = 795) THEN
   		COP(N23[TMP_dSourceOffset], N795[TMP_dDestOffset], TMP_dNumValues);
   	ELSIF (TMP_dSourceFile = 23) AND (TMP_dDestFile = 796) THEN
   		COP(N23[TMP_dSourceOffset], N796[TMP_dDestOffset], TMP_dNumValues);
   	ELSIF (TMP_dSourceFile = 23) AND (TMP_dDestFile = 797) THEN
   		COP(N23[TMP_dSourceOffset], N797[TMP_dDestOffset], TMP_dNumValues);
   	ELSIF (TMP_dSourceFile = 23) AND (TMP_dDestFile = 798) THEN
   		COP(N23[TMP_dSourceOffset], N798[TMP_dDestOffset], TMP_dNumValues);